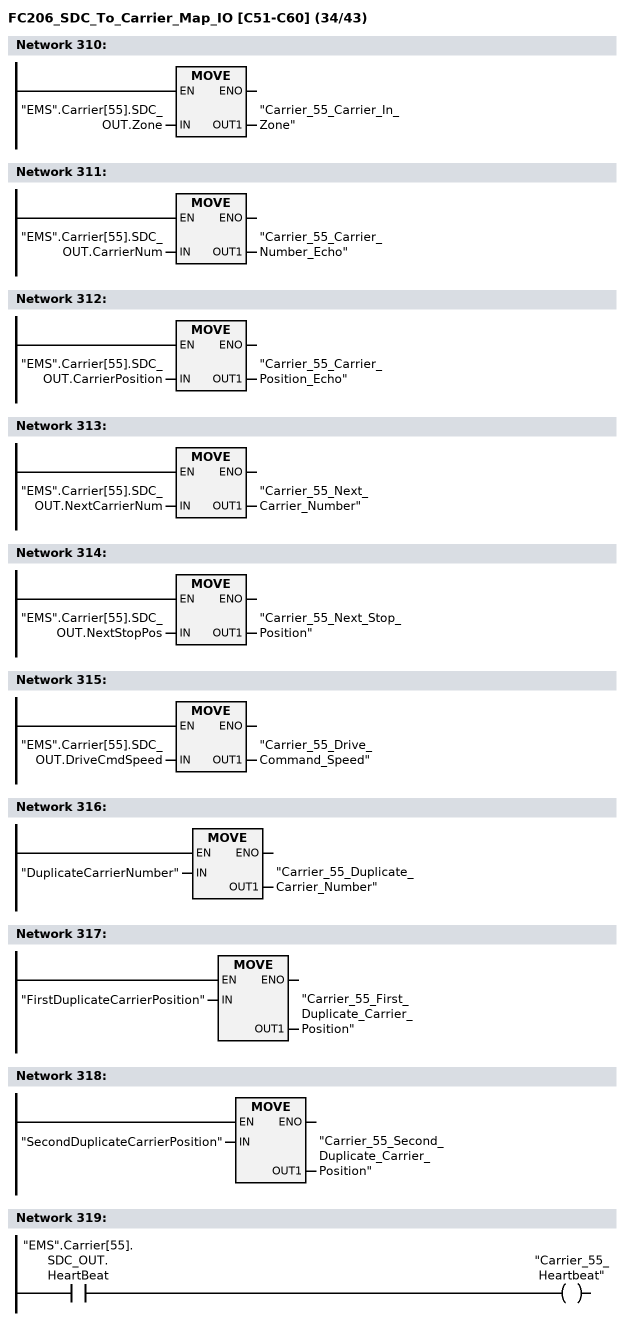
   RUNG wire#powerrail
      Move(in := "EMS".Carrier[55].SDC_OUT.Zone, out1 => "Carrier_55_Carrier_In_Zone")
   END_RUNG
   // the same network as SCL:
   "Carrier_55_Carrier_In_Zone" := "EMS".Carrier[55].SDC_OUT.Zone;
END_REGION

REGION Network 311
   RUNG wire#powerrail
      Move(in := "EMS".Carrier[55].SDC_OUT.CarrierNum, out1 => "Carrier_55_Carrier_Number_Echo")
   END_RUNG
   // the same network as SCL:
   "Carrier_55_Carrier_Number_Echo" := "EMS".Carrier[55].SDC_OUT.CarrierNum;
END_REGION

REGION Network 312
   RUNG wire#powerrail
      Move(in := "EMS".Carrier[55].SDC_OUT.CarrierPosition, out1 => "Carrier_55_Carrier_Position_Echo")
   END_RUNG
   // the same network as SCL:
   "Carrier_55_Carrier_Position_Echo" := "EMS".Carrier[55].SDC_OUT.CarrierPosition;
END_REGION

REGION Network 313
   RUNG wire#powerrail
      Move(in := "EMS".Carrier[55].SDC_OUT.NextCarrierNum, out1 => "Carrier_55_Next_Carrier_Number")
   END_RUNG
   // the same network as SCL:
   "Carrier_55_Next_Carrier_Number" := "EMS".Carrier[55].SDC_OUT.NextCarrierNum;
END_REGION

REGION Network 314
   RUNG wire#powerrail
      Move(in := "EMS".Carrier[55].SDC_OUT.NextStopPos, out1 => "Carrier_55_Next_Stop_Position")
   END_RUNG
   // the same network as SCL:
   "Carrier_55_Next_Stop_Position" := "EMS".Carrier[55].SDC_OUT.NextStopPos;
END_REGION

REGION Network 315
   RUNG wire#powerrail
      Move(in := "EMS".Carrier[55].SDC_OUT.DriveCmdSpeed, out1 => "Carrier_55_Drive_Command_Speed")
   END_RUNG
   // the same network as SCL:
   "Carrier_55_Drive_Command_Speed" := "EMS".Carrier[55].SDC_OUT.DriveCmdSpeed;
END_REGION

REGION Network 316
   RUNG wire#powerrail
      Move(in := "DuplicateCarrierNumber", out1 => "Carrier_55_Duplicate_Carrier_Number")
   END_RUNG
   // the same network as SCL:
   "Carrier_55_Duplicate_Carrier_Number" := "DuplicateCarrierNumber";
END_REGION

REGION Network 317
   RUNG wire#powerrail
      Move(in := "FirstDuplicateCarrierPosition", out1 => "Carrier_55_First_Duplicate_Carrier_Position")
   END_RUNG
   // the same network as SCL:
   "Carrier_55_First_Duplicate_Carrier_Position" := "FirstDuplicateCarrierPosition";
END_REGION

REGION Network 318
   RUNG wire#powerrail
      Move(in := "SecondDuplicateCarrierPosition", out1 => "Carrier_55_Second_Duplicate_Carrier_Position")
   END_RUNG
   // the same network as SCL:
   "Carrier_55_Second_Duplicate_Carrier_Position" := "SecondDuplicateCarrierPosition";
END_REGION

REGION Network 319
   RUNG wire#powerrail
      Contact( "EMS".Carrier[55].SDC_OUT.HeartBeat )
      Coil( "Carrier_55_Heartbeat" )
   END_RUNG
   // the same network as SCL:
   "Carrier_55_Heartbeat" := "EMS".Carrier[55].SDC_OUT.HeartBeat;
END_REGION

REGION Network 320
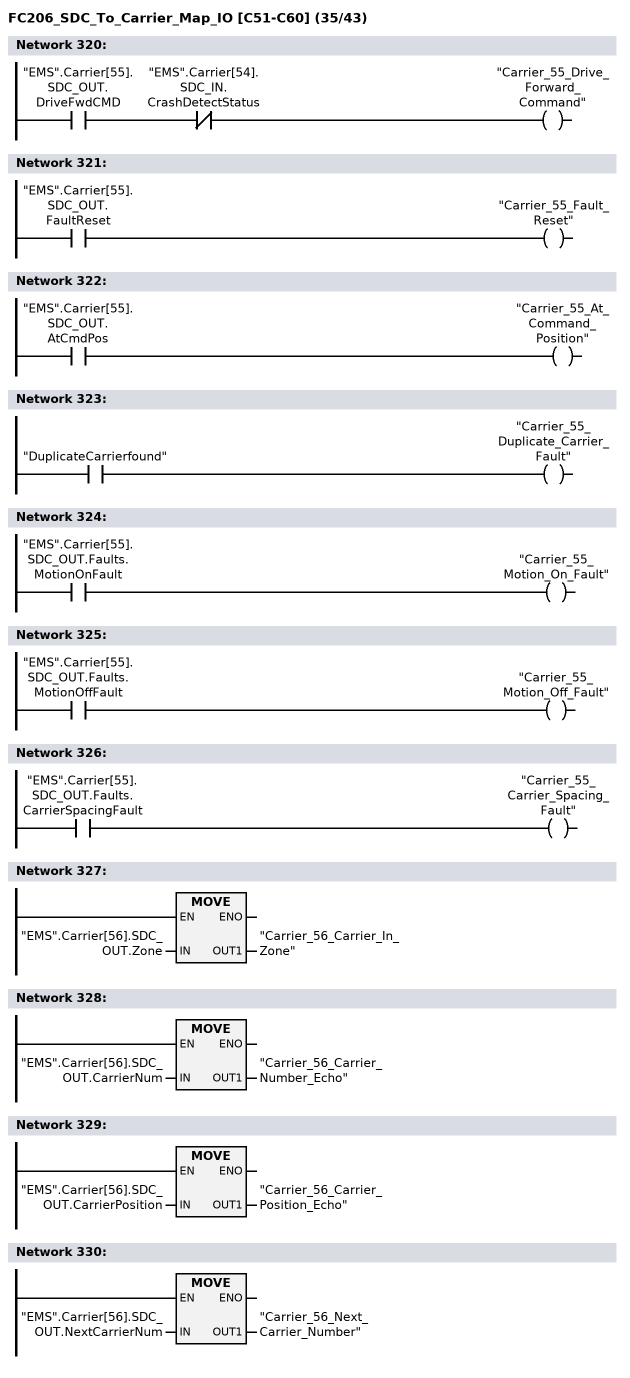
   RUNG wire#powerrail
      Contact( "EMS".Carrier[55].SDC_OUT.DriveFwdCMD )
      I_Contact( "EMS".Carrier[54].SDC_IN.CrashDetectStatus )
      Coil( "Carrier_55_Drive_Forward_Command" )
   END_RUNG
   // the same network as SCL:
   "Carrier_55_Drive_Forward_Command" := "EMS".Carrier[55].SDC_OUT.DriveFwdCMD AND NOT "EMS".Carrier[54].SDC_IN.CrashDetectStatus;
END_REGION

REGION Network 321
   RUNG wire#powerrail
      Contact( "EMS".Carrier[55].SDC_OUT.FaultReset )
      Coil( "Carrier_55_Fault_Reset" )
   END_RUNG
   // the same network as SCL:
   "Carrier_55_Fault_Reset" := "EMS".Carrier[55].SDC_OUT.FaultReset;
END_REGION

REGION Network 322
   RUNG wire#powerrail
      Contact( "EMS".Carrier[55].SDC_OUT.AtCmdPos )
      Coil( "Carrier_55_At_Command_Position" )
   END_RUNG
   // the same network as SCL:
   "Carrier_55_At_Command_Position" := "EMS".Carrier[55].SDC_OUT.AtCmdPos;
END_REGION

REGION Network 323
   RUNG wire#powerrail
      Contact( "DuplicateCarrierfound" )
      Coil( "Carrier_55_Duplicate_Carrier_Fault" )
   END_RUNG
   // the same network as SCL:
   "Carrier_55_Duplicate_Carrier_Fault" := "DuplicateCarrierfound";
END_REGION

REGION Network 324
   RUNG wire#powerrail
      Contact( "EMS".Carrier[55].SDC_OUT.Faults.MotionOnFault )
      Coil( "Carrier_55_Motion_On_Fault" )
   END_RUNG
   // the same network as SCL:
   "Carrier_55_Motion_On_Fault" := "EMS".Carrier[55].SDC_OUT.Faults.MotionOnFault;
END_REGION

REGION Network 325
   RUNG wire#powerrail
      Contact( "EMS".Carrier[55].SDC_OUT.Faults.MotionOffFault )
      Coil( "Carrier_55_Motion_Off_Fault" )
   END_RUNG
   // the same network as SCL:
   "Carrier_55_Motion_Off_Fault" := "EMS".Carrier[55].SDC_OUT.Faults.MotionOffFault;
END_REGION

REGION Network 326
   RUNG wire#powerrail
      Contact( "EMS".Carrier[55].SDC_OUT.Faults.CarrierSpacingFault )
      Coil( "Carrier_55_Carrier_Spacing_Fault" )
   END_RUNG
   // the same network as SCL:
   "Carrier_55_Carrier_Spacing_Fault" := "EMS".Carrier[55].SDC_OUT.Faults.CarrierSpacingFault;
END_REGION

REGION Network 327
   RUNG wire#powerrail
      Move(in := "EMS".Carrier[56].SDC_OUT.Zone, out1 => "Carrier_56_Carrier_In_Zone")
   END_RUNG
   // the same network as SCL:
   "Carrier_56_Carrier_In_Zone" := "EMS".Carrier[56].SDC_OUT.Zone;
END_REGION

REGION Network 328
   RUNG wire#powerrail
      Move(in := "EMS".Carrier[56].SDC_OUT.CarrierNum, out1 => "Carrier_56_Carrier_Number_Echo")
   END_RUNG
   // the same network as SCL:
   "Carrier_56_Carrier_Number_Echo" := "EMS".Carrier[56].SDC_OUT.CarrierNum;
END_REGION

REGION Network 329
   RUNG wire#powerrail
      Move(in := "EMS".Carrier[56].SDC_OUT.CarrierPosition, out1 => "Carrier_56_Carrier_Position_Echo")
   END_RUNG
   // the same network as SCL:
   "Carrier_56_Carrier_Position_Echo" := "EMS".Carrier[56].SDC_OUT.CarrierPosition;
END_REGION

REGION Network 330
   RUNG wire#powerrail
      Move(in := "EMS".Carrier[56].SDC_OUT.NextCarrierNum, out1 => "Carrier_56_Next_Carrier_Number")
   END_RUNG
   // the same network as SCL:
   "Carrier_56_Next_Carrier_Number" := "EMS".Carrier[56].SDC_OUT.NextCarrierNum;
END_REGION

REGION Network 331
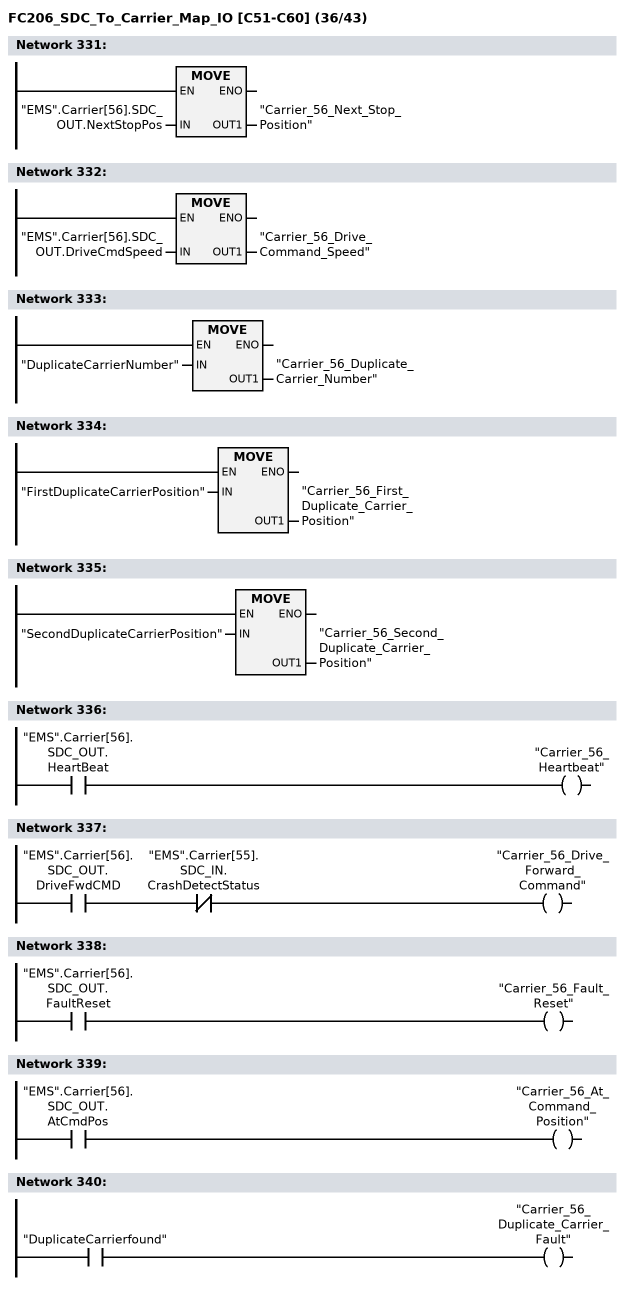
   RUNG wire#powerrail
      Move(in := "EMS".Carrier[56].SDC_OUT.NextStopPos, out1 => "Carrier_56_Next_Stop_Position")
   END_RUNG
   // the same network as SCL:
   "Carrier_56_Next_Stop_Position" := "EMS".Carrier[56].SDC_OUT.NextStopPos;
END_REGION

REGION Network 332
   RUNG wire#powerrail
      Move(in := "EMS".Carrier[56].SDC_OUT.DriveCmdSpeed, out1 => "Carrier_56_Drive_Command_Speed")
   END_RUNG
   // the same network as SCL:
   "Carrier_56_Drive_Command_Speed" := "EMS".Carrier[56].SDC_OUT.DriveCmdSpeed;
END_REGION

REGION Network 333
   RUNG wire#powerrail
      Move(in := "DuplicateCarrierNumber", out1 => "Carrier_56_Duplicate_Carrier_Number")
   END_RUNG
   // the same network as SCL:
   "Carrier_56_Duplicate_Carrier_Number" := "DuplicateCarrierNumber";
END_REGION

REGION Network 334
   RUNG wire#powerrail
      Move(in := "FirstDuplicateCarrierPosition", out1 => "Carrier_56_First_Duplicate_Carrier_Position")
   END_RUNG
   // the same network as SCL:
   "Carrier_56_First_Duplicate_Carrier_Position" := "FirstDuplicateCarrierPosition";
END_REGION

REGION Network 335
   RUNG wire#powerrail
      Move(in := "SecondDuplicateCarrierPosition", out1 => "Carrier_56_Second_Duplicate_Carrier_Position")
   END_RUNG
   // the same network as SCL:
   "Carrier_56_Second_Duplicate_Carrier_Position" := "SecondDuplicateCarrierPosition";
END_REGION

REGION Network 336
   RUNG wire#powerrail
      Contact( "EMS".Carrier[56].SDC_OUT.HeartBeat )
      Coil( "Carrier_56_Heartbeat" )
   END_RUNG
   // the same network as SCL:
   "Carrier_56_Heartbeat" := "EMS".Carrier[56].SDC_OUT.HeartBeat;
END_REGION

REGION Network 337
   RUNG wire#powerrail
      Contact( "EMS".Carrier[56].SDC_OUT.DriveFwdCMD )
      I_Contact( "EMS".Carrier[55].SDC_IN.CrashDetectStatus )
      Coil( "Carrier_56_Drive_Forward_Command" )
   END_RUNG
   // the same network as SCL:
   "Carrier_56_Drive_Forward_Command" := "EMS".Carrier[56].SDC_OUT.DriveFwdCMD AND NOT "EMS".Carrier[55].SDC_IN.CrashDetectStatus;
END_REGION

REGION Network 338
   RUNG wire#powerrail
      Contact( "EMS".Carrier[56].SDC_OUT.FaultReset )
      Coil( "Carrier_56_Fault_Reset" )
   END_RUNG
   // the same network as SCL:
   "Carrier_56_Fault_Reset" := "EMS".Carrier[56].SDC_OUT.FaultReset;
END_REGION

REGION Network 339
   RUNG wire#powerrail
      Contact( "EMS".Carrier[56].SDC_OUT.AtCmdPos )
      Coil( "Carrier_56_At_Command_Position" )
   END_RUNG
   // the same network as SCL:
   "Carrier_56_At_Command_Position" := "EMS".Carrier[56].SDC_OUT.AtCmdPos;
END_REGION

REGION Network 340
   RUNG wire#powerrail
      Contact( "DuplicateCarrierfound" )
      Coil( "Carrier_56_Duplicate_Carrier_Fault" )
   END_RUNG
   // the same network as SCL:
   "Carrier_56_Duplicate_Carrier_Fault" := "DuplicateCarrierfound";
END_REGION

REGION Network 341
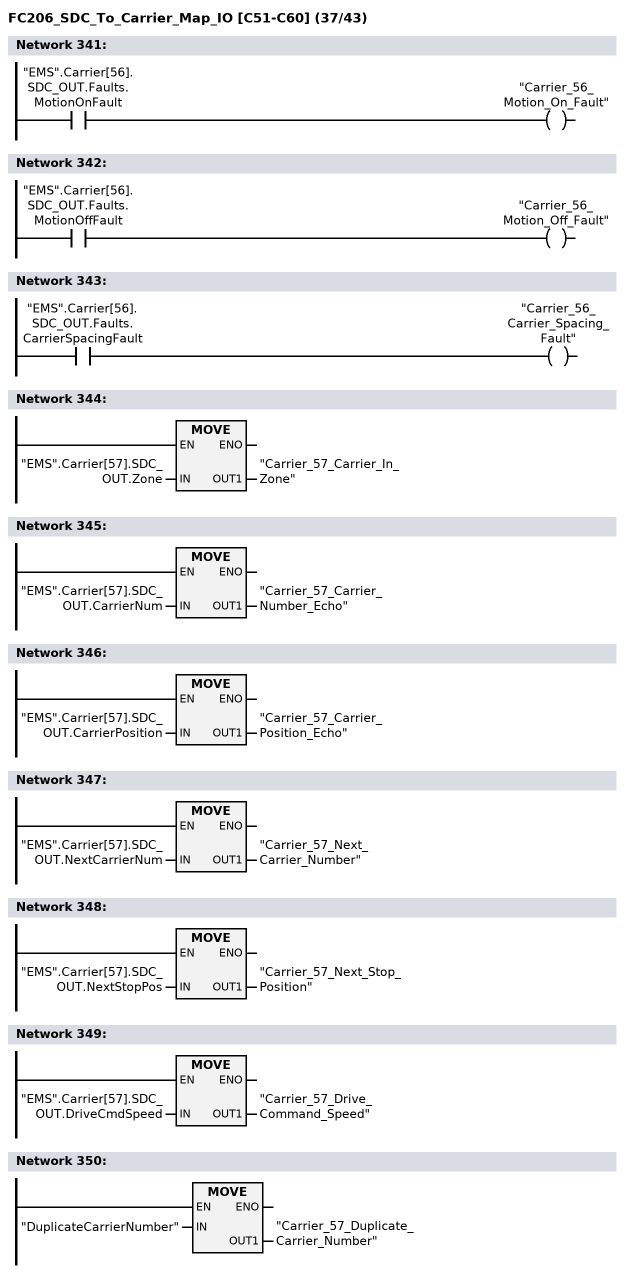
   RUNG wire#powerrail
      Contact( "EMS".Carrier[56].SDC_OUT.Faults.MotionOnFault )
      Coil( "Carrier_56_Motion_On_Fault" )
   END_RUNG
   // the same network as SCL:
   "Carrier_56_Motion_On_Fault" := "EMS".Carrier[56].SDC_OUT.Faults.MotionOnFault;
END_REGION

REGION Network 342
   RUNG wire#powerrail
      Contact( "EMS".Carrier[56].SDC_OUT.Faults.MotionOffFault )
      Coil( "Carrier_56_Motion_Off_Fault" )
   END_RUNG
   // the same network as SCL:
   "Carrier_56_Motion_Off_Fault" := "EMS".Carrier[56].SDC_OUT.Faults.MotionOffFault;
END_REGION

REGION Network 343
   RUNG wire#powerrail
      Contact( "EMS".Carrier[56].SDC_OUT.Faults.CarrierSpacingFault )
      Coil( "Carrier_56_Carrier_Spacing_Fault" )
   END_RUNG
   // the same network as SCL:
   "Carrier_56_Carrier_Spacing_Fault" := "EMS".Carrier[56].SDC_OUT.Faults.CarrierSpacingFault;
END_REGION

REGION Network 344
   RUNG wire#powerrail
      Move(in := "EMS".Carrier[57].SDC_OUT.Zone, out1 => "Carrier_57_Carrier_In_Zone")
   END_RUNG
   // the same network as SCL:
   "Carrier_57_Carrier_In_Zone" := "EMS".Carrier[57].SDC_OUT.Zone;
END_REGION

REGION Network 345
   RUNG wire#powerrail
      Move(in := "EMS".Carrier[57].SDC_OUT.CarrierNum, out1 => "Carrier_57_Carrier_Number_Echo")
   END_RUNG
   // the same network as SCL:
   "Carrier_57_Carrier_Number_Echo" := "EMS".Carrier[57].SDC_OUT.CarrierNum;
END_REGION

REGION Network 346
   RUNG wire#powerrail
      Move(in := "EMS".Carrier[57].SDC_OUT.CarrierPosition, out1 => "Carrier_57_Carrier_Position_Echo")
   END_RUNG
   // the same network as SCL:
   "Carrier_57_Carrier_Position_Echo" := "EMS".Carrier[57].SDC_OUT.CarrierPosition;
END_REGION

REGION Network 347
   RUNG wire#powerrail
      Move(in := "EMS".Carrier[57].SDC_OUT.NextCarrierNum, out1 => "Carrier_57_Next_Carrier_Number")
   END_RUNG
   // the same network as SCL:
   "Carrier_57_Next_Carrier_Number" := "EMS".Carrier[57].SDC_OUT.NextCarrierNum;
END_REGION

REGION Network 348
   RUNG wire#powerrail
      Move(in := "EMS".Carrier[57].SDC_OUT.NextStopPos, out1 => "Carrier_57_Next_Stop_Position")
   END_RUNG
   // the same network as SCL:
   "Carrier_57_Next_Stop_Position" := "EMS".Carrier[57].SDC_OUT.NextStopPos;
END_REGION

REGION Network 349
   RUNG wire#powerrail
      Move(in := "EMS".Carrier[57].SDC_OUT.DriveCmdSpeed, out1 => "Carrier_57_Drive_Command_Speed")
   END_RUNG
   // the same network as SCL:
   "Carrier_57_Drive_Command_Speed" := "EMS".Carrier[57].SDC_OUT.DriveCmdSpeed;
END_REGION

REGION Network 350
   RUNG wire#powerrail
      Move(in := "DuplicateCarrierNumber", out1 => "Carrier_57_Duplicate_Carrier_Number")
   END_RUNG
   // the same network as SCL:
   "Carrier_57_Duplicate_Carrier_Number" := "DuplicateCarrierNumber";
END_REGION

REGION Network 351
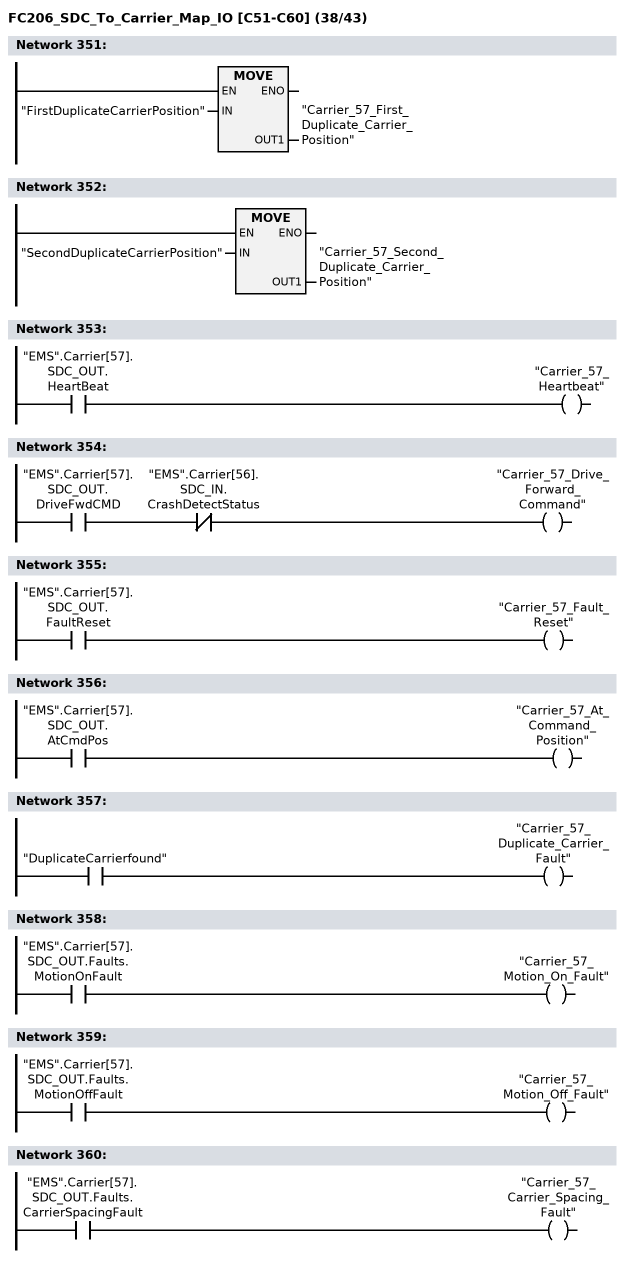
   RUNG wire#powerrail
      Move(in := "FirstDuplicateCarrierPosition", out1 => "Carrier_57_First_Duplicate_Carrier_Position")
   END_RUNG
   // the same network as SCL:
   "Carrier_57_First_Duplicate_Carrier_Position" := "FirstDuplicateCarrierPosition";
END_REGION

REGION Network 352
   RUNG wire#powerrail
      Move(in := "SecondDuplicateCarrierPosition", out1 => "Carrier_57_Second_Duplicate_Carrier_Position")
   END_RUNG
   // the same network as SCL:
   "Carrier_57_Second_Duplicate_Carrier_Position" := "SecondDuplicateCarrierPosition";
END_REGION

REGION Network 353
   RUNG wire#powerrail
      Contact( "EMS".Carrier[57].SDC_OUT.HeartBeat )
      Coil( "Carrier_57_Heartbeat" )
   END_RUNG
   // the same network as SCL:
   "Carrier_57_Heartbeat" := "EMS".Carrier[57].SDC_OUT.HeartBeat;
END_REGION

REGION Network 354
   RUNG wire#powerrail
      Contact( "EMS".Carrier[57].SDC_OUT.DriveFwdCMD )
      I_Contact( "EMS".Carrier[56].SDC_IN.CrashDetectStatus )
      Coil( "Carrier_57_Drive_Forward_Command" )
   END_RUNG
   // the same network as SCL:
   "Carrier_57_Drive_Forward_Command" := "EMS".Carrier[57].SDC_OUT.DriveFwdCMD AND NOT "EMS".Carrier[56].SDC_IN.CrashDetectStatus;
END_REGION

REGION Network 355
   RUNG wire#powerrail
      Contact( "EMS".Carrier[57].SDC_OUT.FaultReset )
      Coil( "Carrier_57_Fault_Reset" )
   END_RUNG
   // the same network as SCL:
   "Carrier_57_Fault_Reset" := "EMS".Carrier[57].SDC_OUT.FaultReset;
END_REGION

REGION Network 356
   RUNG wire#powerrail
      Contact( "EMS".Carrier[57].SDC_OUT.AtCmdPos )
      Coil( "Carrier_57_At_Command_Position" )
   END_RUNG
   // the same network as SCL:
   "Carrier_57_At_Command_Position" := "EMS".Carrier[57].SDC_OUT.AtCmdPos;
END_REGION

REGION Network 357
   RUNG wire#powerrail
      Contact( "DuplicateCarrierfound" )
      Coil( "Carrier_57_Duplicate_Carrier_Fault" )
   END_RUNG
   // the same network as SCL:
   "Carrier_57_Duplicate_Carrier_Fault" := "DuplicateCarrierfound";
END_REGION

REGION Network 358
   RUNG wire#powerrail
      Contact( "EMS".Carrier[57].SDC_OUT.Faults.MotionOnFault )
      Coil( "Carrier_57_Motion_On_Fault" )
   END_RUNG
   // the same network as SCL:
   "Carrier_57_Motion_On_Fault" := "EMS".Carrier[57].SDC_OUT.Faults.MotionOnFault;
END_REGION

REGION Network 359
   RUNG wire#powerrail
      Contact( "EMS".Carrier[57].SDC_OUT.Faults.MotionOffFault )
      Coil( "Carrier_57_Motion_Off_Fault" )
   END_RUNG
   // the same network as SCL:
   "Carrier_57_Motion_Off_Fault" := "EMS".Carrier[57].SDC_OUT.Faults.MotionOffFault;
END_REGION

REGION Network 360
   RUNG wire#powerrail
      Contact( "EMS".Carrier[57].SDC_OUT.Faults.CarrierSpacingFault )
      Coil( "Carrier_57_Carrier_Spacing_Fault" )
   END_RUNG
   // the same network as SCL:
   "Carrier_57_Carrier_Spacing_Fault" := "EMS".Carrier[57].SDC_OUT.Faults.CarrierSpacingFault;
END_REGION

REGION Network 361
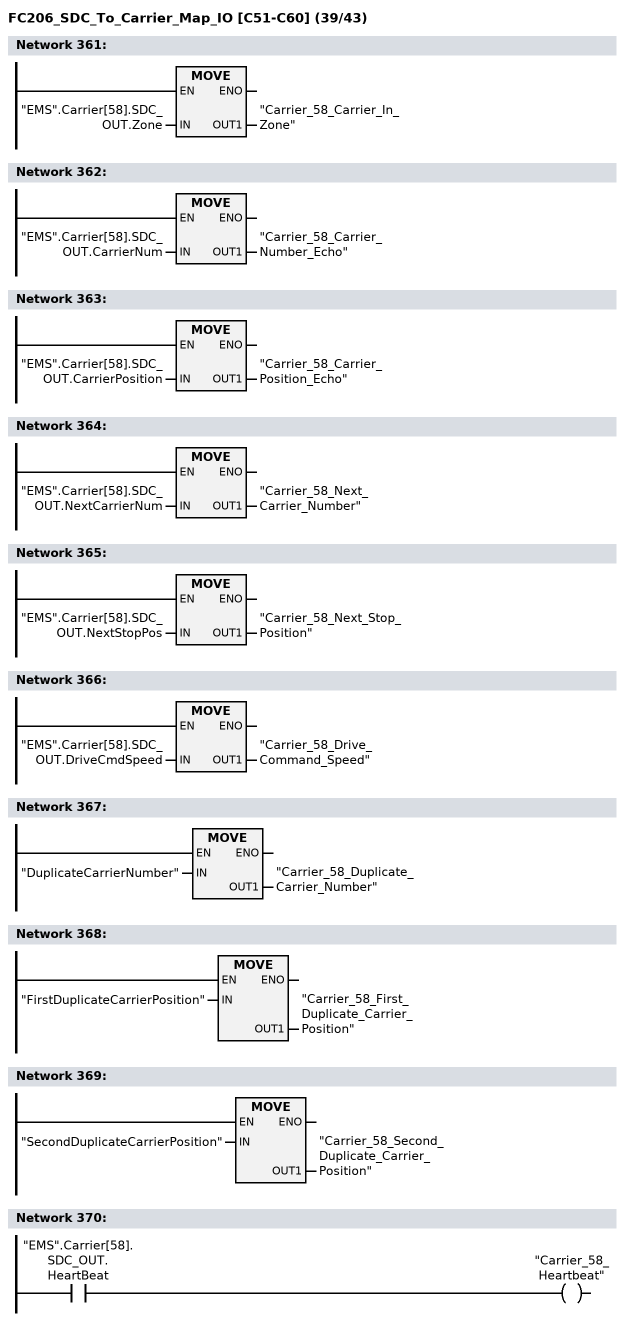
   RUNG wire#powerrail
      Move(in := "EMS".Carrier[58].SDC_OUT.Zone, out1 => "Carrier_58_Carrier_In_Zone")
   END_RUNG
   // the same network as SCL:
   "Carrier_58_Carrier_In_Zone" := "EMS".Carrier[58].SDC_OUT.Zone;
END_REGION

REGION Network 362
   RUNG wire#powerrail
      Move(in := "EMS".Carrier[58].SDC_OUT.CarrierNum, out1 => "Carrier_58_Carrier_Number_Echo")
   END_RUNG
   // the same network as SCL:
   "Carrier_58_Carrier_Number_Echo" := "EMS".Carrier[58].SDC_OUT.CarrierNum;
END_REGION

REGION Network 363
   RUNG wire#powerrail
      Move(in := "EMS".Carrier[58].SDC_OUT.CarrierPosition, out1 => "Carrier_58_Carrier_Position_Echo")
   END_RUNG
   // the same network as SCL:
   "Carrier_58_Carrier_Position_Echo" := "EMS".Carrier[58].SDC_OUT.CarrierPosition;
END_REGION

REGION Network 364
   RUNG wire#powerrail
      Move(in := "EMS".Carrier[58].SDC_OUT.NextCarrierNum, out1 => "Carrier_58_Next_Carrier_Number")
   END_RUNG
   // the same network as SCL:
   "Carrier_58_Next_Carrier_Number" := "EMS".Carrier[58].SDC_OUT.NextCarrierNum;
END_REGION

REGION Network 365
   RUNG wire#powerrail
      Move(in := "EMS".Carrier[58].SDC_OUT.NextStopPos, out1 => "Carrier_58_Next_Stop_Position")
   END_RUNG
   // the same network as SCL:
   "Carrier_58_Next_Stop_Position" := "EMS".Carrier[58].SDC_OUT.NextStopPos;
END_REGION

REGION Network 366
   RUNG wire#powerrail
      Move(in := "EMS".Carrier[58].SDC_OUT.DriveCmdSpeed, out1 => "Carrier_58_Drive_Command_Speed")
   END_RUNG
   // the same network as SCL:
   "Carrier_58_Drive_Command_Speed" := "EMS".Carrier[58].SDC_OUT.DriveCmdSpeed;
END_REGION

REGION Network 367
   RUNG wire#powerrail
      Move(in := "DuplicateCarrierNumber", out1 => "Carrier_58_Duplicate_Carrier_Number")
   END_RUNG
   // the same network as SCL:
   "Carrier_58_Duplicate_Carrier_Number" := "DuplicateCarrierNumber";
END_REGION

REGION Network 368
   RUNG wire#powerrail
      Move(in := "FirstDuplicateCarrierPosition", out1 => "Carrier_58_First_Duplicate_Carrier_Position")
   END_RUNG
   // the same network as SCL:
   "Carrier_58_First_Duplicate_Carrier_Position" := "FirstDuplicateCarrierPosition";
END_REGION

REGION Network 369
   RUNG wire#powerrail
      Move(in := "SecondDuplicateCarrierPosition", out1 => "Carrier_58_Second_Duplicate_Carrier_Position")
   END_RUNG
   // the same network as SCL:
   "Carrier_58_Second_Duplicate_Carrier_Position" := "SecondDuplicateCarrierPosition";
END_REGION

REGION Network 370
   RUNG wire#powerrail
      Contact( "EMS".Carrier[58].SDC_OUT.HeartBeat )
      Coil( "Carrier_58_Heartbeat" )
   END_RUNG
   // the same network as SCL:
   "Carrier_58_Heartbeat" := "EMS".Carrier[58].SDC_OUT.HeartBeat;
END_REGION

REGION Network 371
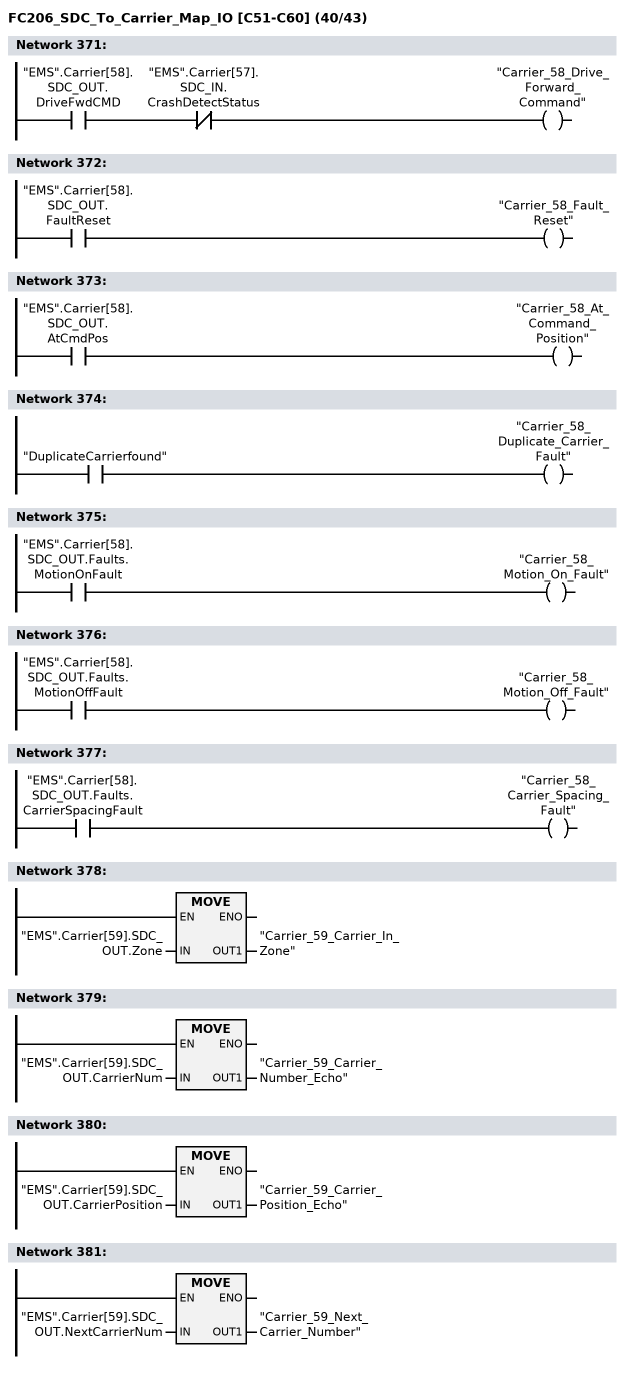
   RUNG wire#powerrail
      Contact( "EMS".Carrier[58].SDC_OUT.DriveFwdCMD )
      I_Contact( "EMS".Carrier[57].SDC_IN.CrashDetectStatus )
      Coil( "Carrier_58_Drive_Forward_Command" )
   END_RUNG
   // the same network as SCL:
   "Carrier_58_Drive_Forward_Command" := "EMS".Carrier[58].SDC_OUT.DriveFwdCMD AND NOT "EMS".Carrier[57].SDC_IN.CrashDetectStatus;
END_REGION

REGION Network 372
   RUNG wire#powerrail
      Contact( "EMS".Carrier[58].SDC_OUT.FaultReset )
      Coil( "Carrier_58_Fault_Reset" )
   END_RUNG
   // the same network as SCL:
   "Carrier_58_Fault_Reset" := "EMS".Carrier[58].SDC_OUT.FaultReset;
END_REGION

REGION Network 373
   RUNG wire#powerrail
      Contact( "EMS".Carrier[58].SDC_OUT.AtCmdPos )
      Coil( "Carrier_58_At_Command_Position" )
   END_RUNG
   // the same network as SCL:
   "Carrier_58_At_Command_Position" := "EMS".Carrier[58].SDC_OUT.AtCmdPos;
END_REGION

REGION Network 374
   RUNG wire#powerrail
      Contact( "DuplicateCarrierfound" )
      Coil( "Carrier_58_Duplicate_Carrier_Fault" )
   END_RUNG
   // the same network as SCL:
   "Carrier_58_Duplicate_Carrier_Fault" := "DuplicateCarrierfound";
END_REGION

REGION Network 375
   RUNG wire#powerrail
      Contact( "EMS".Carrier[58].SDC_OUT.Faults.MotionOnFault )
      Coil( "Carrier_58_Motion_On_Fault" )
   END_RUNG
   // the same network as SCL:
   "Carrier_58_Motion_On_Fault" := "EMS".Carrier[58].SDC_OUT.Faults.MotionOnFault;
END_REGION

REGION Network 376
   RUNG wire#powerrail
      Contact( "EMS".Carrier[58].SDC_OUT.Faults.MotionOffFault )
      Coil( "Carrier_58_Motion_Off_Fault" )
   END_RUNG
   // the same network as SCL:
   "Carrier_58_Motion_Off_Fault" := "EMS".Carrier[58].SDC_OUT.Faults.MotionOffFault;
END_REGION

REGION Network 377
   RUNG wire#powerrail
      Contact( "EMS".Carrier[58].SDC_OUT.Faults.CarrierSpacingFault )
      Coil( "Carrier_58_Carrier_Spacing_Fault" )
   END_RUNG
   // the same network as SCL:
   "Carrier_58_Carrier_Spacing_Fault" := "EMS".Carrier[58].SDC_OUT.Faults.CarrierSpacingFault;
END_REGION

REGION Network 378
   RUNG wire#powerrail
      Move(in := "EMS".Carrier[59].SDC_OUT.Zone, out1 => "Carrier_59_Carrier_In_Zone")
   END_RUNG
   // the same network as SCL:
   "Carrier_59_Carrier_In_Zone" := "EMS".Carrier[59].SDC_OUT.Zone;
END_REGION

REGION Network 379
   RUNG wire#powerrail
      Move(in := "EMS".Carrier[59].SDC_OUT.CarrierNum, out1 => "Carrier_59_Carrier_Number_Echo")
   END_RUNG
   // the same network as SCL:
   "Carrier_59_Carrier_Number_Echo" := "EMS".Carrier[59].SDC_OUT.CarrierNum;
END_REGION

REGION Network 380
   RUNG wire#powerrail
      Move(in := "EMS".Carrier[59].SDC_OUT.CarrierPosition, out1 => "Carrier_59_Carrier_Position_Echo")
   END_RUNG
   // the same network as SCL:
   "Carrier_59_Carrier_Position_Echo" := "EMS".Carrier[59].SDC_OUT.CarrierPosition;
END_REGION

REGION Network 381
   RUNG wire#powerrail
      Move(in := "EMS".Carrier[59].SDC_OUT.NextCarrierNum, out1 => "Carrier_59_Next_Carrier_Number")
   END_RUNG
   // the same network as SCL:
   "Carrier_59_Next_Carrier_Number" := "EMS".Carrier[59].SDC_OUT.NextCarrierNum;
END_REGION

REGION Network 382
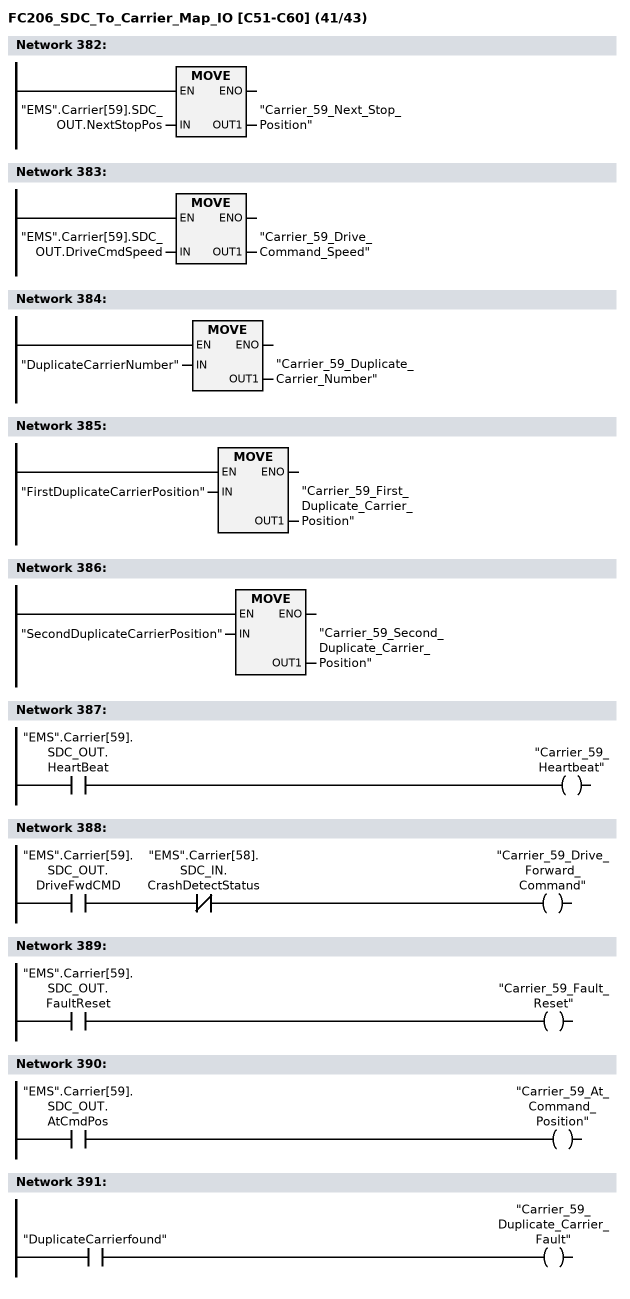
   RUNG wire#powerrail
      Move(in := "EMS".Carrier[59].SDC_OUT.NextStopPos, out1 => "Carrier_59_Next_Stop_Position")
   END_RUNG
   // the same network as SCL:
   "Carrier_59_Next_Stop_Position" := "EMS".Carrier[59].SDC_OUT.NextStopPos;
END_REGION

REGION Network 383
   RUNG wire#powerrail
      Move(in := "EMS".Carrier[59].SDC_OUT.DriveCmdSpeed, out1 => "Carrier_59_Drive_Command_Speed")
   END_RUNG
   // the same network as SCL:
   "Carrier_59_Drive_Command_Speed" := "EMS".Carrier[59].SDC_OUT.DriveCmdSpeed;
END_REGION

REGION Network 384
   RUNG wire#powerrail
      Move(in := "DuplicateCarrierNumber", out1 => "Carrier_59_Duplicate_Carrier_Number")
   END_RUNG
   // the same network as SCL:
   "Carrier_59_Duplicate_Carrier_Number" := "DuplicateCarrierNumber";
END_REGION

REGION Network 385
   RUNG wire#powerrail
      Move(in := "FirstDuplicateCarrierPosition", out1 => "Carrier_59_First_Duplicate_Carrier_Position")
   END_RUNG
   // the same network as SCL:
   "Carrier_59_First_Duplicate_Carrier_Position" := "FirstDuplicateCarrierPosition";
END_REGION

REGION Network 386
   RUNG wire#powerrail
      Move(in := "SecondDuplicateCarrierPosition", out1 => "Carrier_59_Second_Duplicate_Carrier_Position")
   END_RUNG
   // the same network as SCL:
   "Carrier_59_Second_Duplicate_Carrier_Position" := "SecondDuplicateCarrierPosition";
END_REGION

REGION Network 387
   RUNG wire#powerrail
      Contact( "EMS".Carrier[59].SDC_OUT.HeartBeat )
      Coil( "Carrier_59_Heartbeat" )
   END_RUNG
   // the same network as SCL:
   "Carrier_59_Heartbeat" := "EMS".Carrier[59].SDC_OUT.HeartBeat;
END_REGION

REGION Network 388
   RUNG wire#powerrail
      Contact( "EMS".Carrier[59].SDC_OUT.DriveFwdCMD )
      I_Contact( "EMS".Carrier[58].SDC_IN.CrashDetectStatus )
      Coil( "Carrier_59_Drive_Forward_Command" )
   END_RUNG
   // the same network as SCL:
   "Carrier_59_Drive_Forward_Command" := "EMS".Carrier[59].SDC_OUT.DriveFwdCMD AND NOT "EMS".Carrier[58].SDC_IN.CrashDetectStatus;
END_REGION

REGION Network 389
   RUNG wire#powerrail
      Contact( "EMS".Carrier[59].SDC_OUT.FaultReset )
      Coil( "Carrier_59_Fault_Reset" )
   END_RUNG
   // the same network as SCL:
   "Carrier_59_Fault_Reset" := "EMS".Carrier[59].SDC_OUT.FaultReset;
END_REGION

REGION Network 390
   RUNG wire#powerrail
      Contact( "EMS".Carrier[59].SDC_OUT.AtCmdPos )
      Coil( "Carrier_59_At_Command_Position" )
   END_RUNG
   // the same network as SCL:
   "Carrier_59_At_Command_Position" := "EMS".Carrier[59].SDC_OUT.AtCmdPos;
END_REGION

REGION Network 391
   RUNG wire#powerrail
      Contact( "DuplicateCarrierfound" )
      Coil( "Carrier_59_Duplicate_Carrier_Fault" )
   END_RUNG
   // the same network as SCL:
   "Carrier_59_Duplicate_Carrier_Fault" := "DuplicateCarrierfound";
END_REGION

REGION Network 392
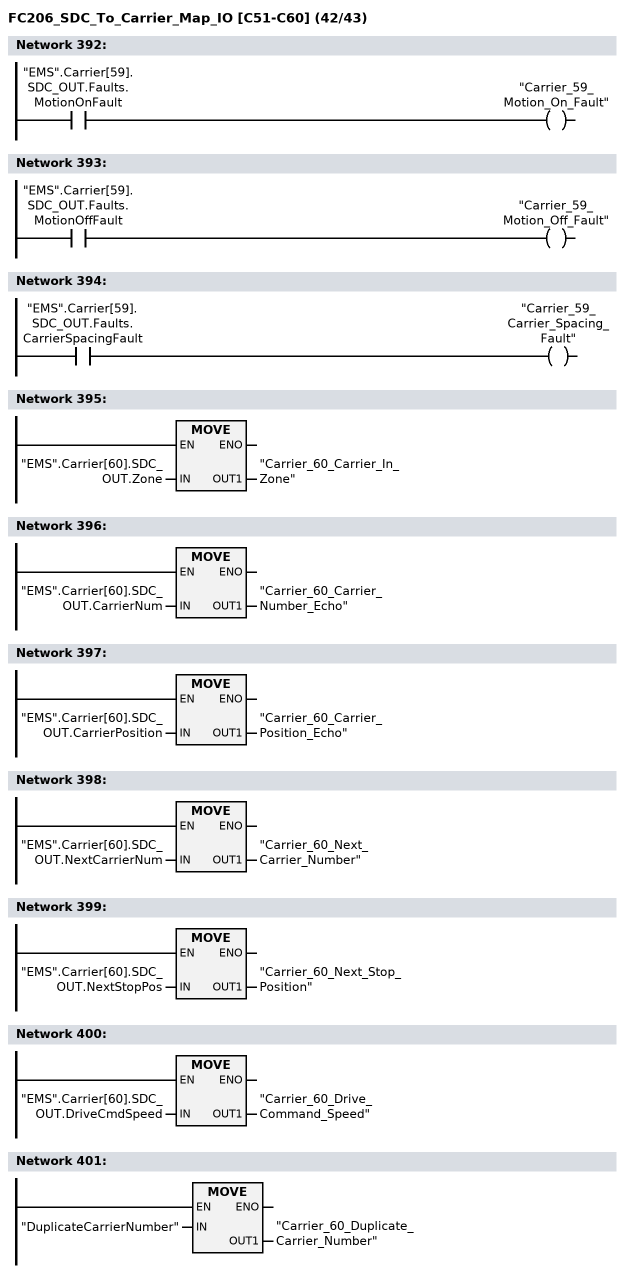
   RUNG wire#powerrail
      Contact( "EMS".Carrier[59].SDC_OUT.Faults.MotionOnFault )
      Coil( "Carrier_59_Motion_On_Fault" )
   END_RUNG
   // the same network as SCL:
   "Carrier_59_Motion_On_Fault" := "EMS".Carrier[59].SDC_OUT.Faults.MotionOnFault;
END_REGION

REGION Network 393
   RUNG wire#powerrail
      Contact( "EMS".Carrier[59].SDC_OUT.Faults.MotionOffFault )
      Coil( "Carrier_59_Motion_Off_Fault" )
   END_RUNG
   // the same network as SCL:
   "Carrier_59_Motion_Off_Fault" := "EMS".Carrier[59].SDC_OUT.Faults.MotionOffFault;
END_REGION
